
                   REGION Program funckji
                       REGION Symulacja wejsc - przepisywanie wartosci wejsciowych, gdy nie ma symulacji oprocz bWeAkt
                           IF "DB352_FF8".FF8[#i].bSt_Tryb.%X12 = 0 THEN
                               "DB352_FF8".FF8[#i].bSym.%X1 := "DB352_FF8".FF8[#i].bWeZalAuto;
                               "DB352_FF8".FF8[#i].bSym.%X8 := "DB352_FF8".FF8[#i].bWeBlZmAuto;
                               "DB352_FF8".FF8[#i].bSym.%X9 := "DB352_FF8".FF8[#i].bWeIlock;
                           END_IF;
                       END_REGION
                       REGION Okreslenie stanow
                           "DB352_FF8".FF8[#i].bSt_Tryb.%X8 := "DB352_FF8".FF8[#i].bWeAkt;
                           "DB352_FF8".FF8[#i].bSt_Tryb.%X9 := (("DB352_FF8".FF8[#i].bSym.%X8 AND "DB352_FF8".FF8[#i].bSt_Tryb.%X12) OR ("DB321_DIO".DIO[#i].bWeBlZmAuto AND NOT "DB352_FF8".FF8[#i].bSt_Tryb.%X12));
                           "DB352_FF8".FF8[#i].bSt_Tryb.%X11 := (("DB352_FF8".FF8[#i].bWeIlock AND NOT "DB352_FF8".FF8[#i].bSt_Tryb.%X12) OR ("DB352_FF8".FF8[#i].bSym.%X9 AND "DB352_FF8".FF8[#i].bSt_Tryb.%X12));
                           "DB352_FF8".FF8[#i].bSt_Tryb.%X12 := "DB352_FF8".FF8[#i].bRoZB1.%X1;
                       END_REGION
                       REGION Licznik czasu trwania impulsu
                           IF "DB352_FF8".FF8[#i].bRoZB1.%X3 AND #Imp_Sek AND NOT "DB352_FF8".FF8[#i].bPauza AND "DB352_FF8".FF8[#i].dT2_Akt=0  THEN
                               CASE "DB352_FF8".FF8[#i].iPetle OF
                                   0: "DB352_FF8".FF8[#i].dT1_old := "DB352_FF8".FF8[#i].dT1i;
                                       GOTO Warunek1;

                                   1: "DB352_FF8".FF8[#i].dT1_old := "DB352_FF8".FF8[#i].dT2i;
                                       GOTO Warunek1;

                                   2: "DB352_FF8".FF8[#i].dT1_old := "DB352_FF8".FF8[#i].dT3i;
                                       GOTO Warunek1;

                                   3: "DB352_FF8".FF8[#i].dT1_old := "DB352_FF8".FF8[#i].dT4i;
                                       GOTO Warunek1;

                                   4: "DB352_FF8".FF8[#i].dT1_old := "DB352_FF8".FF8[#i].dT5i;
                                       GOTO Warunek1;

                                   5: "DB352_FF8".FF8[#i].dT1_old := "DB352_FF8".FF8[#i].dT6i;
                                       GOTO Warunek1;

                                   6: "DB352_FF8".FF8[#i].dT1_old := "DB352_FF8".FF8[#i].dT7i;
                                       GOTO Warunek1;

                                   7: "DB352_FF8".FF8[#i].dT1_old := "DB352_FF8".FF8[#i].dT8i;
                                       GOTO Warunek1;

                                   ELSE
                                       GOTO Warunek1;
                                       ;
                               END_CASE;
                           ELSE
                               GOTO Warunek2;
                               ;
                           END_IF;
                       Warunek1:
                           "DB352_FF8".FF8[#i].dT1_Akt:="DB352_FF8".FF8[#i].dT1_Akt+1;
                           IF "DB352_FF8".FF8[#i].dT1_Akt>="DB352_FF8".FF8[#i].dT1_old THEN
                               "DB352_FF8".FF8[#i].bIhlp := 1;
                               "DB352_FF8".FF8[#i].dT1_Akt := 0;
                               "DB352_FF8".FF8[#i].iPetle := "DB352_FF8".FF8[#i].iPetle + 1;
                               ;
                           END_IF;

                           REGION Ustawianie bitu Pauzy
                           Warunek2:
                               "DB352_FF8".FF8[#i].bPauza:="DB352_FF8".FF8[#i].iPetle>="DB352_FF8".FF8[#i].iIG;
                           END_REGION
                           REGION Licznik czasu trwania przerwy miedzy impulsami
                               IF #Imp_Sek AND "DB352_FF8".FF8[#i].bRoZB1.%X3 AND NOT "DB352_FF8".FF8[#i].bPauza AND "DB352_FF8".FF8[#i].bIhlp  THEN
                                   "DB352_FF8".FF8[#i].dT2_Akt := "DB352_FF8".FF8[#i].dT2_Akt + 1;
                                   IF "DB352_FF8".FF8[#i].dT2_Akt>="DB352_FF8".FF8[#i].dT2 THEN
                                       "DB352_FF8".FF8[#i].bIhlp := 0;
                                       "DB352_FF8".FF8[#i].dT2_Akt := 0;
                                   END_IF;
                               END_IF;
                           END_REGION
                           REGION Licznik czasu trwania przerwy miedzy grupami impulsow
                               IF #Imp_Sek AND "DB352_FF8".FF8[#i].bPauza  THEN
                                   "DB352_FF8".FF8[#i].dT3_Akt := "DB352_FF8".FF8[#i].dT3_Akt + 1;
                                   IF "DB352_FF8".FF8[#i].dT3_Akt>="DB352_FF8".FF8[#i].dT3 THEN
                                       "DB352_FF8".FF8[#i].bIhlp := 0;
                                       "DB352_FF8".FF8[#i].dT3_Akt := 0;
                                       "DB352_FF8".FF8[#i].iPetle := 0;
                                   END_IF;
                               END_IF;
                           END_REGION
                           REGION Wyjscia
                               "DB352_FF8".FF8[#i].bI8 := NOT "DB352_FF8".FF8[#i].bIhlp AND "DB352_FF8".FF8[#i].iPetle = 7;

                               "DB352_FF8".FF8[#i].bI7 := NOT "DB352_FF8".FF8[#i].bIhlp AND "DB352_FF8".FF8[#i].iPetle = 6;

                               "DB352_FF8".FF8[#i].bI6 := NOT "DB352_FF8".FF8[#i].bIhlp AND "DB352_FF8".FF8[#i].iPetle = 5;

                               "DB352_FF8".FF8[#i].bI5 := NOT "DB352_FF8".FF8[#i].bIhlp AND "DB352_FF8".FF8[#i].iPetle = 4;

                               "DB352_FF8".FF8[#i].bI4 := NOT "DB352_FF8".FF8[#i].bIhlp AND "DB352_FF8".FF8[#i].iPetle = 3;

                               "DB352_FF8".FF8[#i].bI3 := NOT "DB352_FF8".FF8[#i].bIhlp AND "DB352_FF8".FF8[#i].iPetle = 2;

                               "DB352_FF8".FF8[#i].bI2 := NOT "DB352_FF8".FF8[#i].bIhlp AND "DB352_FF8".FF8[#i].iPetle = 1;

                               "DB352_FF8".FF8[#i].bI1 := NOT "DB352_FF8".FF8[#i].bIhlp AND "DB352_FF8".FF8[#i].iPetle = 0;
                           END_REGION
                           REGION Wylaczenie
                               IF NOT "DB352_FF8".FF8[#i].bRoZB1.%X3 THEN
                                   "DB352_FF8".FF8[#i].dT1_Akt := 0;
                                   "DB352_FF8".FF8[#i].dT2_Akt := 0;
                                   "DB352_FF8".FF8[#i].dT3_Akt := 0;
                                   "DB352_FF8".FF8[#i].bIhlp := 0;
                                   "DB352_FF8".FF8[#i].bI1 := 0;
                                   "DB352_FF8".FF8[#i].bI2 := 0;
                                   "DB352_FF8".FF8[#i].bI3 := 0;
                                   "DB352_FF8".FF8[#i].bI4 := 0;
                                   "DB352_FF8".FF8[#i].bI5 := 0;
                                   "DB352_FF8".FF8[#i].bI6 := 0;
                                   "DB352_FF8".FF8[#i].bI7 := 0;
                                   "DB352_FF8".FF8[#i].bI8 := 0;
                               END_IF;
                           END_REGION
                       END_REGION
                       REGION Tryb pracy i sterowanie wyjsciem
                           REGION Przepisanie potwierdzen na sterowanie reczne gdy tryb zdalny-auto
                               // Przypadek gdy ktos z wlaczonym lokalnie urz. przechodzi na tryb zdalny-reczny
                               IF "DB352_FF8".FF8[#i].bTrP=8 THEN
                                   "DB352_FF8".FF8[#i].bRoZB1.%X3 := (("DB352_FF8".FF8[#i].bWeZalAuto AND NOT "DB352_FF8".FF8[#i].bSt_Tryb.%X12) OR ("DB352_FF8".FF8[#i].bSym.%X1 AND "DB352_FF8".FF8[#i].bSt_Tryb.%X12));
                               END_IF;

                           END_REGION

                           REGION Blokada zmiany trybu zdalny-automatyczny
                               IF (("DB352_FF8".FF8[#i].bWeBlZmAuto AND NOT "DB352_FF8".FF8[#i].bSt_Tryb.%X12) OR ("DB352_FF8".FF8[#i].bSym.%X8 AND "DB352_FF8".FF8[#i].bSt_Tryb.%X12)) AND "DB352_FF8".FF8[#i].bTrP.%X3 THEN
                                   "DB352_FF8".FF8[#i].bRoZB1.%X0 := 1;
                               END_IF;
                           END_REGION
                           REGION Okreslenie trybu pracy wyjscia
                               IF "DB352_FF8".FF8[#i].bRoZB1.%X0 AND NOT "DB352_FF8".FF8[#i].bSt_Tryb.%X9 THEN
                                   "DB352_FF8".FF8[#i].bTrP := 8;
                               END_IF;
                               IF NOT "DB352_FF8".FF8[#i].bRoZB1.%X0 THEN
                                   "DB352_FF8".FF8[#i].bTrP := 4
                                   ;
                               END_IF;
                           END_REGION
                           REGION Sterowanie wyjsciem
                               "DB352_FF8".FF8[#i].bWySter := "DB352_FF8".FF8[#i].bWeZalAuto;
                           END_REGION
                           REGION Stan urzadzenia
                               IF "DB352_FF8".FF8[#i].bWySter THEN
                                   "DB352_FF8".FF8[#i].bSt_Urz := 8; //urz. wlaczone
                               ELSE
                                   "DB352_FF8".FF8[#i].bSt_Urz := 8; //urz. wylaczone
                               END_IF;
                           END_REGION
                       END_REGION
                       REGION Ustawienia koncowe
                           // Samokasowanie sygnalow
                           IF "DB352_FF8".FF8[#i].bAoff = 1 THEN
                               "DB352_FF8".FF8[#i].bWeZalAuto := 0;
                           END_IF;
                       END_REGION
                   END_REGION
               END_IF;
          END_REGION
     END_FOR;
END_FUNCTION

FUNCTION "FC353_TMR" : Void   // FC353, SCL
{ S7_Optimized_Access := 'TRUE' }
VERSION : 0.1
   VAR_INPUT
      Nr_Ost_Elementu : Int;
      Nr_Plc : Byte;
   END_VAR
   VAR_TEMP
      i : Int;
      TmrTyp : Int;
   END_VAR
BEGIN

   FOR #i := 1 TO #Nr_Ost_Elementu BY 1 DO
       REGION Opisy bitow sygnalow: bRoz,bSym,bSt,bSt_1,bTrP

           //bRoz - ROZKAZ OPERATORA - DB353.DBW10 - WORD
           //bRozB1
           //"DB353_TMR".TMR[#i].bRoZB1.%X0 - Tryb pracy: 0-Zdalny reczny; 1-Zdalny auto
           //"DB353_TMR".TMR[#i].bRoZB1.%X1 - Symulacja wejsc urz: 0-Wylaczona; 1-Zalaczona
           //"DB353_TMR".TMR[#i].bRoZB1.%X2 - Rezerwa
           //"DB353_TMR".TMR[#i].bRoZB1.%X3 - Sterowanie urz. w tr. Zdalnym-Man: 0-Wylacz; 1-Zalacz
           //"DB353_TMR".TMR[#i].bRoZB1.%X4-X7 - Rezerwa
           //
           //bRozB2 - impulsy
           //"DB353_TMR".TMR[#i].bRoZB2.%X0-X7 - Rezerwa (impuls)
           //
           //bSym - SYM WEJSCIA - DB353.DBW12 - WORD
           //"DB353_TMR".TMR[#i].bSym.%X0 - Aktywacja urz. w systemie (ustawiany tylko z programu)
           //"DB353_TMR".TMR[#i].bSym.%X1 - Sterowanie urz. w tr. Zdalnym-Auto: 0-Wylacz; 1-Zalacz
           //"DB353_TMR".TMR[#i].bSym.%X2-X7 - Rezerwa
           //"DB353_TMR".TMR[#i].bSym.%X8 - Blokada zmiany tr. zdalnego z Auto na Man: 0-Brak; 1-Aktywna
           //"DB353_TMR".TMR[#i].bSym.%X9 - Interlock w trybie Zdalnym-Auto: 0-Brak; 1-Aktywny
           //"DB353_TMR".TMR[#i].bSym.%X10-X11 - Rezerwa
           //"DB353_TMR".TMR[#i].bSym.%X12 - Zerowanie timera (kasowanie przez obiekt)
           //"DB353_TMR".TMR[#i].bSym.%X13-X15 - Rezerwa
           //
           //bSt_Tryb - STAN - DB353.DBW14 - WORD
           //"DB353_TMR".TMR[#i].bSt_Tryb.%X0-X7
           //"DB353_TMR".TMR[#i].bSt_Tryb.%X8 - Urzadzenie aktywowane
           //"DB353_TMR".TMR[#i].bSt_Tryb.%X9 - Blokada zmaiany tr. zdalnego z Auto na Man: 0-Brak; 1-Aktywna
           //"DB353_TMR".TMR[#i].bSt_Tryb.%X10 - Stan rezerwa
           //"DB353_TMR".TMR[#i].bSt_Tryb.%X11 - Interlock w trybie Zdalnym-Auto: 0-Brak; 1-Aktywny
           //"DB353_TMR".TMR[#i].bSt_Tryb.%X12 - Symulacja wejsc urzadzenia: 0-Wylaczona; 1-Zalaczona
           //"DB353_TMR".TMR[#i].bSt_Tryb.%X13 - Rezerwa
           //"DB353_TMR".TMR[#i].bSt_Tryb.%X14 - Rezerwa
           //"DB353_TMR".TMR[#i].bSt_Tryb.%X15 - Rezerwa
           //
           //bSt_Urz - STAN - DB353.DBW16 - INT
           //"DB353_TMR".TMR[#i].bSt_Urz.%X0 - STAN(1)- Awaria zbiorcza 1-Aktywna; 0-Brak aktywnosci obiektu
           //"DB353_TMR".TMR[#i].bSt_Urz.%X1 - STAN(2)- Urzadzenie: 1-Zamkniete; 0-Inny stan
           //"DB353_TMR".TMR[#i].bSt_Urz.%X2 - STAN(4)- Rezerwa
           //"DB353_TMR".TMR[#i].bSt_Urz.%X3 - STAN(8)- Urzadzenie: 1-Otwarte; 0-Inny stan
           //"DB353_TMR".TMR[#i].bSt_Urz.%X4 - STAN(16)- Rezerwa
           //"DB353_TMR".TMR[#i].bSt_Urz.%X5 - STAN(32)- Rezerwa
           //"DB353_TMR".TMR[#i].bSt_Urz.%X6-X7 - STAN(64)(128)- Rezerwa
           //
           //bTrP - TRYB PRACY - DB353.DBW17 - INT
           //"DB353_TMR".TMR[#i].bTrP.%X0 - TRYB PRACY(1) - Rezerwa
           //"DB353_TMR".TMR[#i].bTrP.%X1 - Tryb PRACY(2) - Rezerwa
           //"DB353_TMR".TMR[#i].bTrP.%X2 - TRYB PRACY(4) - Tryb Sterowania Zdalnego: 1-Zdalny Reczny; 0-Inny stan
           //"DB353_TMR".TMR[#i].bTrP.%X3 - TRYB PRACY(8) - Tryb Sterowania Zdalnego: 1-Zdalny Automatyczny; 0-Inny stan
           //"DB353_TMR".TMR[#i].bTrP.%X4-X7 - Tryb PRACY(16)(32)(64)(128) - Rezerwa
       END_REGION
       REGION Przepisanie danych do obiektu
           "DB353_TMR".TMR[#i].yNrID := #i;
           "DB353_TMR".TMR[#i].yNrPLC := #Nr_Plc;
       END_REGION
       REGION Warunek na wykonanie funkcji
           IF "DB353_TMR".TMR[#i].bWeAkt = 0 THEN //Akcja przy deaktywowaniu obiektu
               "DB353_TMR".TMR[#i].bWeAkt := 0;
               "DB353_TMR".TMR[#i].bWeZalAuto := 0;
               "DB353_TMR".TMR[#i].bWeBlZmAuto := 0;
               "DB353_TMR".TMR[#i].bWeIlock := 0;
               "DB353_TMR".TMR[#i].bWeZeruj := 0;
               "DB353_TMR".TMR[#i].bRoZB1 := 0;
               "DB353_TMR".TMR[#i].bSym := 0;
               "DB353_TMR".TMR[#i].bSt_Tryb := 0;
               "DB353_TMR".TMR[#i].bSt_Urz := 0;
               "DB353_TMR".TMR[#i].bTrP := 0;
               "DB353_TMR".TMR[#i].bWySter := 0;
           ELSE

               REGION Program funckji
                   REGION Symulacja wejsc - przepisywanie wartosci wejsciowych, gdy nie ma symulacji oprocz bWeAkt
                       IF "DB353_TMR".TMR[#i].bSt_Tryb.%X12 = 0 THEN
                           "DB353_TMR".TMR[#i].bSym.%X1 := "DB353_TMR".TMR[#i].bWeZalAuto;
                           "DB353_TMR".TMR[#i].bSym.%X8 := "DB353_TMR".TMR[#i].bWeBlZmAuto;
                           "DB353_TMR".TMR[#i].bSym.%X9 := "DB353_TMR".TMR[#i].bWeIlock;
                           "DB353_TMR".TMR[#i].bSym.%X12 := "DB353_TMR".TMR[#i].bWeZeruj;
                       END_IF;
                   END_REGION
                   REGION Okreslenie stanow
                       "DB353_TMR".TMR[#i].bSt_Tryb.%X8 := "DB353_TMR".TMR[#i].bWeAkt;
                       "DB353_TMR".TMR[#i].bSt_Tryb.%X9 := (("DB353_TMR".TMR[#i].bSym.%X8 AND "DB353_TMR".TMR[#i].bSt_Tryb.%X12) OR ("DB353_TMR".TMR[#i].bWeBlZmAuto AND NOT "DB353_TMR".TMR[#i].bSt_Tryb.%X12));
                       "DB353_TMR".TMR[#i].bSt_Tryb.%X11 := (("DB353_TMR".TMR[#i].bWeIlock AND NOT "DB353_TMR".TMR[#i].bSt_Tryb.%X12) OR ("DB353_TMR".TMR[#i].bSym.%X9 AND "DB353_TMR".TMR[#i].bSt_Tryb.%X12));
                       "DB353_TMR".TMR[#i].bSt_Tryb.%X12 := "DB353_TMR".TMR[#i].bRoZB1.%X1;
                   END_REGION
                   REGION Licznik czasu
                           IF "DB353_TMR".TMR[#i].bLatch THEN
                               #TmrTyp := 5;
                           ELSE
                               #TmrTyp := 1;
                           END_IF;

                           IF NOT "DB353_TMR".TMR[#i].bSt_Tryb.%X11 THEN
                               "FC301_Timer"(iTyp := #TmrTyp,
                                             bOnOff := ("DB353_TMR".TMR[#i].bSym.%X1 AND "DB353_TMR".TMR[#i].bSt_Tryb.%X12) OR ("DB353_TMR".TMR[#i].bWeZalAuto AND NOT "DB353_TMR".TMR[#i].bSt_Tryb.%X12),
                                             bRst := ("DB353_TMR".TMR[#i].bSym.%X12 AND "DB353_TMR".TMR[#i].bSt_Tryb.%X12) OR ("DB353_TMR".TMR[#i].bWeZeruj AND NOT "DB353_TMR".TMR[#i].bSt_Tryb.%X12),
                                             dCzasZad := "DB353_TMR".TMR[#i].dCzZad,
                                             timer_1s := "imp1s",
                                             bOk => "DB353_TMR".TMR[#i].bHlp187,
                                             dCzasAkt := "DB353_TMR".TMR[#i].dCzAkt);

                           END_IF;


                   END_REGION
                   REGION Tryb pracy i sterowanie wyjsciem
                       REGION Przepisanie potwierdzen na sterowanie reczne gdy tryb zdalny-auto
                           // Przypadek gdy ktos z wlaczonym lokalnie urz. przechodzi na tryb zdalny-reczny
                           IF "DB353_TMR".TMR[#i].bTrP = 8 THEN
                               "DB353_TMR".TMR[#i].bRoZB1.%X3 := (("DB353_TMR".TMR[#i].bWeZalAuto AND NOT "DB353_TMR".TMR[#i].bSt_Tryb.%X12) OR ("DB353_TMR".TMR[#i].bSym.%X1 AND "DB353_TMR".TMR[#i].bSt_Tryb.%X12));
                           END_IF;

                       END_REGION

                       REGION Blokada zmiany trybu zdalny-automatyczny
                           IF (("DB353_TMR".TMR[#i].bWeBlZmAuto AND NOT "DB353_TMR".TMR[#i].bSt_Tryb.%X12) OR ("DB353_TMR".TMR[#i].bSym.%X8 AND "DB353_TMR".TMR[#i].bSt_Tryb.%X12)) AND "DB353_TMR".TMR[#i].bTrP.%X3 THEN
                               "DB353_TMR".TMR[#i].bRoZB1.%X0 := 1;
                           END_IF;
                       END_REGION
                       REGION Okreslenie trybu pracy wyjscia
                           IF "DB353_TMR".TMR[#i].bRoZB1.%X0 AND NOT "DB353_TMR".TMR[#i].bSt_Tryb.%X9 THEN
                               "DB353_TMR".TMR[#i].bTrP := 8;
                           END_IF;
                           IF NOT "DB353_TMR".TMR[#i].bRoZB1.%X0 THEN
                               "DB353_TMR".TMR[#i].bTrP := 4
                               ;
                           END_IF;
                       END_REGION
                       REGION Sterowanie wyjsciem
                           "DB353_TMR".TMR[#i].bWySter := "DB353_TMR".TMR[#i].bHlp187;
                       END_REGION
                       REGION Stan urzadzenia
                           IF (("DB353_TMR".TMR[#i].bSym.%X1 AND "DB353_TMR".TMR[#i].bSt_Tryb.%X12) OR ("DB353_TMR".TMR[#i].bWeZalAuto AND NOT "DB353_TMR".TMR[#i].bSt_Tryb.%X12)) OR "DB353_TMR".TMR[#i].bWySter THEN
                               "DB353_TMR".TMR[#i].bSt_Urz := 8; //urz. wlaczone
                           ELSE
                               "DB353_TMR".TMR[#i].bSt_Urz := 2; //urz. wylaczone
                           END_IF;
                       END_REGION
                   END_REGION
                   REGION Ustawienia koncowe
                       // Samokasowanie sygnalow

                       IF ("DB353_TMR".TMR[#i].bSym.%X12 AND "DB353_TMR".TMR[#i].bSt_Tryb.%X12) OR ("DB353_TMR".TMR[#i].bWeZeruj AND NOT "DB353_TMR".TMR[#i].bSt_Tryb.%X12) THEN
                           "DB353_TMR".TMR[#i].bSym.%X12 := 0;
                           "DB353_TMR".TMR[#i].bWeZeruj := 0;
                       END_IF;

                       IF "DB353_TMR".TMR[#i].bAoff = 1 THEN
                           "DB353_TMR".TMR[#i].bWeZalAuto := 0;
                       END_IF;

                   END_REGION
               END_REGION
           END_IF;
       END_REGION
   END_FOR;
END_FUNCTION

FUNCTION "FC1000_System" : Void   // FC1000, LAD
{ S7_Optimized_Access := 'TRUE' }
VERSION : 0.1
   VAR_TEMP   // added for the SCL form of the ladder/FBD networks
      _w1 : Bool;
   END_VAR
BEGIN

REGION Network 1: Imp 1s
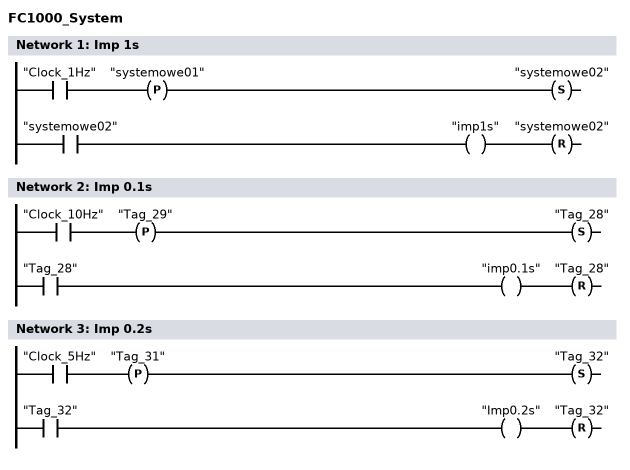
   RUNG wire#powerrail
      Contact( "Clock_1Hz" )
      P_Trig( "systemowe01" )
      S_Coil( "systemowe02" )
   END_RUNG
   RUNG wire#powerrail
      Contact( "systemowe02" )
      Coil( "imp1s" )
      R_Coil( "systemowe02" )
   END_RUNG
   // the same network as SCL:
   #_w1 := "Clock_1Hz" AND NOT "systemowe01";   // rising edge
   "systemowe01" := "Clock_1Hz";
   IF #_w1 THEN "systemowe02" := TRUE; END_IF;
   "imp1s" := "systemowe02";
   IF "systemowe02" THEN "systemowe02" := FALSE; END_IF;
END_REGION

REGION Network 2: Imp 0.1s
   RUNG wire#powerrail
      Contact( "Clock_10Hz" )
      P_Trig( "Tag_29" )
      S_Coil( "Tag_28" )
   END_RUNG
   RUNG wire#powerrail
      Contact( "Tag_28" )
      Coil( "imp0.1s" )
      R_Coil( "Tag_28" )
   END_RUNG
   // the same network as SCL:
   #_w1 := "Clock_10Hz" AND NOT "Tag_29";   // rising edge
   "Tag_29" := "Clock_10Hz";
   IF #_w1 THEN "Tag_28" := TRUE; END_IF;
   "imp0.1s" := "Tag_28";
   IF "Tag_28" THEN "Tag_28" := FALSE; END_IF;
END_REGION

REGION Network 3: Imp 0.2s
   RUNG wire#powerrail
      Contact( "Clock_5Hz" )
      P_Trig( "Tag_31" )
      S_Coil( "Tag_32" )
   END_RUNG
   RUNG wire#powerrail
      Contact( "Tag_32" )
      Coil( "Imp0.2s" )
      R_Coil( "Tag_32" )
   END_RUNG
   // the same network as SCL:
   #_w1 := "Clock_5Hz" AND NOT "Tag_31";   // rising edge
   "Tag_31" := "Clock_5Hz";
   IF #_w1 THEN "Tag_32" := TRUE; END_IF;
   "Imp0.2s" := "Tag_32";
   IF "Tag_32" THEN "Tag_32" := FALSE; END_IF;
END_REGION
END_FUNCTION

// folder: Sinamics

FUNCTION_BLOCK "DM_Objects"   // FB1, LAD
{ S7_Optimized_Access := 'TRUE' }
VERSION : 0.1
   VAR
      pump1Tank1out : "DM_Class";
      pump2Tank1in : "DM_Class";
   END_VAR
   VAR_TEMP
      i : Int;
   END_VAR
BEGIN

REGION Network 1 (SCL): Wpisanie parametrow
   #pump2Tank1in.inCircBreaker := true;
   #pump2Tank1in.inPTC := TRUE;

   #pump1Tank1out.inCircBreaker := true;
   #pump1Tank1out.inPTC := TRUE;
END_REGION

REGION Network 2: Wywolanie obiektu LAD
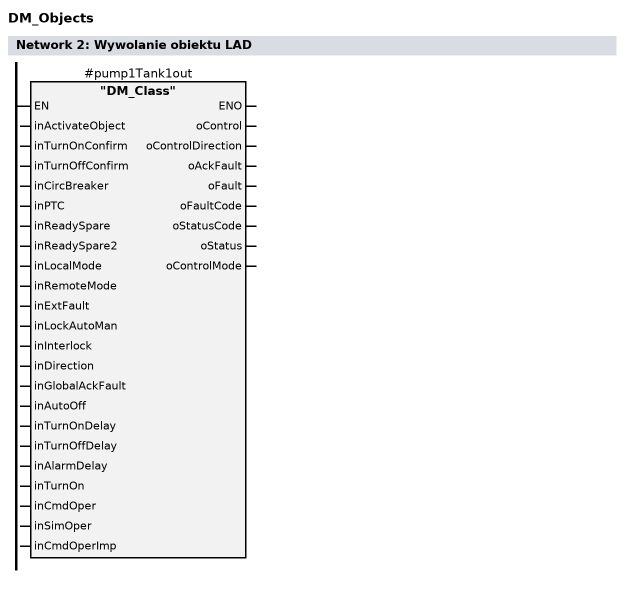
   RUNG wire#powerrail
      #pump1Tank1out(inActivateObject :=, inTurnOnConfirm :=, inTurnOffConfirm :=, inCircBreaker :=, inPTC :=, inReadySpare :=, inReadySpare2 :=, inLocalMode :=, inRemoteMode :=, inExtFault :=, inLockAutoMan :=, inInterlock :=, inDirection :=, inGlobalAckFault :=, inAutoOff :=, inTurnOnDelay :=, inTurnOffDelay :=, inAlarmDelay :=, inTurnOn :=, inCmdOper :=, inSimOper :=, inCmdOperImp :=, oControl =>, oControlDirection =>, oAckFault =>, oFault =>, oFaultCode =>, oStatusCode =>, oStatus =>, oControlMode =>)
   END_RUNG
   // the same network as SCL:
   #pump1Tank1out();   // "DM_Class"
END_REGION

REGION Network 3 (SCL): Wywolanie obiektu SCL - ladniejsze
   #pump2Tank1in();
END_REGION
END_FUNCTION_BLOCK

FUNCTION_BLOCK "DM_Sinamics"   // FB2, SCL
{ S7_Optimized_Access := 'TRUE' }
VERSION : 0.1
   VAR
      pump1Power : MC_POWER;
      pump1Control : MC_MOVEJOG;
      pump2Power : MC_POWER;
      pump2Control : MC_MOVEJOG;
   END_VAR
BEGIN

   REGION Pump 1

       #pump1Power(Axis:="pump1",
                   Enable:=NOT "DB_DM".pump1Tank1out.oFault);

       #pump1Control(Axis := "pump2",
                     JogForward := "DB_DM".pump1Tank1out.oControl AND NOT "DB_DM".pump1Tank1out.oControlDirection,
                     JogBackward := "DB_DM".pump1Tank1out.oControl AND "DB_DM".pump1Tank1out.oControlDirection);

   END_REGION


   REGION Pump 2

       #pump2Power(Axis := "pump2",
                   Enable := NOT "DB_DM".pump2Tank1in.oFault);

       #pump2Control(Axis := "pump2",
                     JogForward := "DB_DM".pump2Tank1in.oControl AND NOT "DB_DM".pump2Tank1in.oControlDirection,
                     JogBackward := "DB_DM".pump2Tank1in.oControl AND "DB_DM".pump2Tank1in.oControlDirection);

   END_REGION
END_FUNCTION_BLOCK

FUNCTION_BLOCK "DM_Class"   // FB301, SCL
{ S7_Optimized_Access := 'TRUE' }
VERSION : 0.1
   VAR_INPUT
      inActivateObject : Bool := true;   // Aktywowanie działania obiektu
      inTurnOnConfirm : Bool;   // Potwierdzenie załączenia
      inTurnOffConfirm : Bool;   // Potwierdzenie wyłączenia
      inCircBreaker : Bool;   // Gotowość obiektu - rozłącznik
      inPTC : Bool;   // Gotowość obiektu - PTC
      inReadySpare : Bool := true;   // Gotowość obiektu - rezerwa
      inReadySpare2 : Bool := true;   // Gotowość obiektu - rezerwa
      inLocalMode : Bool;   // Tryb lokalny
      inRemoteMode : Bool;   // Tryb remontowy
      inExtFault : Bool;   // Błąd zewnętrzny
      inLockAutoMan : Bool;   // Blokada przełączenia trybu Auto-Manual
      inInterlock : Bool;   // Interlok
      inDirection : Bool;   // Kierunek obrotów (1-odwrotny)
      inGlobalAckFault : Bool;   // Globalny reset
      inAutoOff : Bool;   // Resetowanie sterowania na końcu
      inTurnOnDelay : DInt;   // Czas opóźnienia załączenia [s]
      inTurnOffDelay : DInt;   // Czas opóźnienia wyłączenia [s]
      inAlarmDelay : DInt;   // Czas opóźnienia alarmu od potwierdzeń [s]
   END_VAR
   VAR_OUTPUT
      oControl : Bool;   // Wyjście sterujące
      oControlDirection : Bool;   // Wyjście strujące kierunkiem obrotów
      oAckFault : Bool;   // Wyjście reset obiektu
      oFault : Bool;   // Wyjście awaria
      oFaultCode : Byte;   // Kod awarii
      oStatusCode : Word;   // Kod statusu
      oStatus : Int;   // Status ( 1-awaria; 2-Wył; 4-Załączanie; 8-Zał; 16-Wyłączanie)
      oControlMode : Int;   // Tryb pracy (1-remont; 2-lokal; 4-manual; 8-auto)
   END_VAR
   VAR_IN_OUT
      inTurnOn : Bool;   // Załączanie z programu
      inCmdOper : Word := 16#5;   // Komendy manualne
      inSimOper : Word;   // Komendy symulacji
      inCmdOperImp : Word;   // Komendy impulsowe
   END_VAR
   VAR
      statReady : Bool;
      statManAuto : Bool;
      statSymOn : Bool;
      statSwitchEnable : Bool;
      statManTurnOn : Bool;
      statManDirection : Bool;
      statSwitchControl : Bool;
      statFaultReset : Bool;
      statActivate : Bool;
      statTurnOn : Bool;
      statTurnOnConfirm : Bool;
      statTurnOffConfirm : Bool;
      statLocal : Bool;
      statRemote : Bool;
      statExtFault : Bool;
      statLockAutoMan : Bool;
      statInterlock : Bool;
      statDirection : Bool;
      tofTurnOnDelay : TON_TIME;
      tofTurnOffDelay : TOF_TIME;
      tonAlarm : TON_TIME;
      statAlarmStart : Bool;
      statFault : Bool;
      statControlMode : Int;
      statControl : Bool;
      statTmrOnOff : Bool;
      trigGlobalReset : R_TRIG;
   END_VAR
BEGIN
   REGION Activation object - condition to execute function
       IF NOT #inActivateObject THEN
           #inTurnOn := FALSE;
           #inCmdOper := 0;
           #inSimOper := 0;
           #inCmdOperImp := 0;

           #oControl := FALSE;
           #oControlDirection := FALSE;
           #oAckFault := FALSE;
           #oFault := FALSE;
           #oFaultCode := 0;
           #oStatusCode := 0;
           #oStatus := 0;
           #oControlMode := 0;

           RETURN;

       END_IF;

   END_REGION

   REGION Rewriting inputs

       //Operator Control Word
       #statManAuto := #inCmdOper.%X0;
       #statSymOn := #inCmdOper.%X1;
       #statSwitchEnable := #inCmdOper.%X2;
       #statManTurnOn := #inCmdOper.%X3;
       #statManDirection := #inCmdOper.%X4;
       #statSwitchControl := #inCmdOper.%X6;

       //Operator Control Word Impulses
       #trigGlobalReset(CLK:=#inGlobalAckFault);

       #statFaultReset := #trigGlobalReset.Q OR #inCmdOperImp.%X0;

   END_REGION

   REGION Rewriting inputs or simulation signals to statics

       IF NOT #statSymOn THEN

           #statTurnOn := #inTurnOn;
           #statTurnOnConfirm := #inTurnOnConfirm;
           #statTurnOffConfirm := #inTurnOffConfirm;
           #statReady := #inCircBreaker AND #inPTC AND #inReadySpare AND #inReadySpare2 ;
           #statLocal := #inLocalMode;
           #statRemote := #inRemoteMode;
           #statExtFault := #inExtFault;
           #statLockAutoMan := #inLockAutoMan;
           #statInterlock := #inInterlock;
           #statDirection := #inDirection;

           //Rewriting inputs to simulation bits when simulotion is to switch fluently
           #inSimOper.%X0 := #statActivate;
           #inSimOper.%X1 := #statTurnOn;
           #inSimOper.%X2 := #statTurnOnConfirm;
           #inSimOper.%X3 := #statTurnOffConfirm;
           #inSimOper.%X4 := #statReady;
           #inSimOper.%X5 := #statLocal;
           #inSimOper.%X6 := #statRemote;
           #inSimOper.%X7 := #statExtFault;
           #inSimOper.%X8 := #statLockAutoMan;
           #inSimOper.%X9 := #statInterlock;
           #inSimOper.%X10 := #statDirection;

       ELSE

           #statActivate := #inSimOper.%X0;
           #statTurnOn := #inSimOper.%X1;
           #statTurnOnConfirm := #inSimOper.%X2;
           #statTurnOffConfirm := #inSimOper.%X3;
           #statReady:= #inSimOper.%X4;
           #statLocal := #inSimOper.%X5;
           #statRemote := #inSimOper.%X6;
           #statExtFault := #inSimOper.%X7;
           #statLockAutoMan := #inSimOper.%X8;
           #statInterlock := #inSimOper.%X9;
           #statDirection := #inSimOper.%X10;

       END_IF;


   END_REGION

   REGION Control Mode

       IF #statRemote THEN

           #statControlMode := 1;

       ELSIF #statLocal THEN

           #statControlMode := 2;

       ELSIF NOT #statManAuto AND NOT #statLockAutoMan THEN

           #statControlMode := 4;

       ELSIF #statManAuto AND NOT #statLockAutoMan THEN

           #statControlMode := 8;

       END_IF;

   END_REGION

   REGION TurnOn/Off Delay

       #tofTurnOnDelay(IN := #statTurnOn,
                       PT := 1000 * #inTurnOnDelay);

       #tofTurnOffDelay(IN := #statTurnOn,
                        PT := 1000 * #inTurnOffDelay);

       IF #tofTurnOnDelay.Q THEN

           #statTmrOnOff := TRUE;

       END_IF;

       IF NOT #tofTurnOffDelay.Q THEN

           #statTmrOnOff := FALSE;

       END_IF;
   END_REGION

   REGION Fault 
       //Zerowanie czasu awari przy zmianie sterowanie podczas ruchu - czy to w ogole cokolwiek robi???

       //Alarm from switching control 
       #statAlarmStart :=
       #statSwitchControl AND //is switch controling on
       #statSwitchEnable AND //is objects output is eneble to turn on
       #statControlMode<>2 AND //in local mode there is no alarm
       #statControlMode<>1 AND //in remote mode there is no alarm
       (
       (#statControl XOR #statTurnOnConfirm) OR //xor  0110 - if A and B have different state then =1
       (NOT #statControl XOR #statTurnOffConfirm) OR
       (#statTurnOnConfirm AND #statTurnOffConfirm) OR
       (NOT #statTurnOnConfirm AND NOT #statTurnOffConfirm)
       )
       ;
       //#tonAlarm.PT := DINT_TO_TIME(1000 * #AlarmDelay);
       //Generating switching alarm after delay
       #tonAlarm(IN := #statAlarmStart,
                 PT:=DINT_TO_TIME(1000 * #inAlarmDelay));


       //Generating fault
       IF #tonAlarm.Q OR NOT #statReady OR #statExtFault THEN

           #statFault := TRUE;

       ELSIF #statFaultReset THEN

           #statFault := FALSE;

       END_IF;

       //Fault reset 
       // IF #statFaultReset THEN
       //     #statFault := FALSE;


       // END_IF;

       //Fault code
       #oFaultCode.%X0 := #tonAlarm.Q;
       #oFaultCode.%X1 := NOT #statReady;
       #oFaultCode.%X2 := #statExtFault;
       #oFaultCode.%X3 := NOT #inCircBreaker;
       #oFaultCode.%X4 := NOT #inPTC;
       #oFaultCode.%X5 := NOT #inReadySpare;
       #oFaultCode.%X6 := NOT #inReadySpare2;

   END_REGION

   REGION Command locks

       IF #statControlMode = 8 AND #statLockAutoMan THEN

           #statManAuto := TRUE;

       ELSIF #statControlMode = 4 AND #statLockAutoMan THEN

           #statManAuto := FALSE;

       END_IF;

       // Writing states from Local to Manual when object when switching Local to Manual
       IF #statControlMode = 2 THEN

           #statManAuto := FALSE;

           IF #statTurnOffConfirm THEN

               #statTurnOn := FALSE;

           ELSIF #statTurnOnConfirm THEN

               #statTurnOn := TRUE;

           END_IF;

       END_IF;

       // Writing states from Auto to Manual when object when switching Auto to Manual
       // Przypadek gdy ktos z wlaczonym automatycznie urz. przechodzi na tryb zdalny-reczny
       IF #statControlMode = 8 THEN

           #statManTurnOn := #statTurnOn;
           #statManDirection := #statDirection;

       END_IF;

       //Resetowanie rozkazu zalaczenia w trybie manualnym po awarii
       IF #statFault THEN

           #statManTurnOn := FALSE;

       END_IF;




   END_REGION

   REGION Control output

       #statControl :=
       #statSwitchEnable AND
       NOT #statInterlock AND
       NOT #statFault AND
       ((#statControlMode = 8 AND #statTmrOnOff) OR
       (#statControlMode = 4 AND #statManTurnOn));

   END_REGION

   REGION Control Direction Output

       #oControlDirection :=
       #statSwitchEnable AND
       ((#statControlMode = 8 AND #statDirection) OR
       (#statControlMode = 4 AND #statManDirection));

   END_REGION

   REGION Reset Control

       #oAckFault := #statFaultReset;

   END_REGION ;

   REGION Device status code
       IF #statFault THEN
           #oStatus := 1;

       ELSIF #statControlMode = 1 THEN
           #oStatus := 2;

       ELSIF #statControlMode = 2 THEN

           IF #statTurnOnConfirm THEN
               #oStatus := 8;

           ELSIF #statTurnOffConfirm THEN
               #oStatus := 2;

           ELSIF #statControl THEN
               #oStatus := 4;

           ELSIF NOT #statControl THEN
               #oStatus := 16;
           END_IF;

       ELSIF #statControlMode > 2 THEN

           IF #statSwitchControl AND #statSwitchEnable THEN

               IF #statControl AND NOT #statTurnOffConfirm AND #statTurnOnConfirm THEN

                   #oStatus := 8;

               ELSIF NOT #statControl AND NOT #statTurnOnConfirm AND #statTurnOffConfirm THEN

                   #oStatus := 2;

               ELSIF #statControl THEN

                   #oStatus := 4;

               ELSIF NOT #statControl THEN

                   #oStatus := 16;

               END_IF;

           ELSIF NOT #statSwitchControl OR NOT #statSwitchEnable THEN //if no output enable or switch check then

               IF #statControl THEN

                   #oStatus := 8;

               ELSIF NOT #statControl THEN

                   #oStatus := 2;

               END_IF;

           END_IF;

       ELSE
           #oStatus := 0;

       END_IF;

   END_REGION ;


   REGION Reseting impuls
       // Samokasowanie sygnalow
       #statFaultReset := false;

       IF #inAutoOff THEN

           #statTurnOn := FALSE;

       END_IF;

   END_REGION ;

   REGION Status code


   END_REGION

   REGION Rewriting TO outputs

       #inCmdOper.%X0 := #statManAuto;
       #inCmdOper.%X1 := #statSymOn;
       #inCmdOper.%X2 := #statSwitchEnable;
       #inCmdOper.%X3 := #statManTurnOn;
       #inCmdOper.%X4 := #statManDirection;
       #inCmdOper.%X6 := #statSwitchControl;

       #inCmdOperImp.%X0 := #statFaultReset;

       #oControlMode := #statControlMode;

       #oFault := #statFault;

       #inTurnOn := #statTurnOn;

       #oControl := #statControl;
   END_REGION
END_FUNCTION_BLOCK

// ===== library types =====

// folder: LGF/4 Math operations

FUNCTION_BLOCK "LGF_Integration"   // FB10043, SCL
TITLE = LGF_Integration
{ S7_Optimized_Access := 'TRUE' }
AUTHOR : Siemens_Digital_Industries
FAMILY : LGF
NAME : LGF_Integration
// The function approximately calculates the area under a function curve. The function curve is transferred as an analog `value` (LReal) which varies over time. The integral value is output on `integral`.  
// The implementation is based on the trapezoidal rule and uses [ms] as time base.
// Diese Funktion  berechnet näherungsweise die Fläche unter einer Funktionskurve. Die Funktionskurve wird als Analogwert `value` (LReal) übergeben, der über die Zeit variiert. Am Ausgang  `integral`wird der Integralwert ausgegeben.  
// Die Implementierung beruht auf der Trapetzmethode und nutzt [ms] als Zeitbasis.
   VAR_INPUT
      enable : Bool;   // Enables integral calculation If this input is set to the value `FALSE`, the integral calculation is stopped and the `integral` output shows the last calculated value. / Aktivierung der Integral Rechnung Wird dieser Eingang auf den Wert `FALSE` berechnung gestoppt und der Ausgang `integral` zeigt den zuletzt berechneten Wert.
      value : LReal;   // Analog value of the continuous function curve, based on [ms], (e.g. [volume flow/ms]) / Analogwert der kontinuierlichen Funktionskurve, basierent auf [ms], (z.B. [Volumenstrom/ms])
      reset : Bool;   // Sets the output “integral” to “0.0”. / Setzt den Ausgang "integral" auf "0.0".
   END_VAR
   VAR_OUTPUT
      integral : LReal;   // Integral value / Integral Wert
      error : Bool;   // FALSE: No error TRUE: An error occurred during the execution of the FB / FALSE: Kein Fehler TRUE: Während der Ausführung des FB ist ein Fehler aufgetreten
      status : Word;   // 16#0000-16#7FFF: Status des FB 16#8000-16#FFFF: Fehleridentifikation (siehe folgende Tabelle) / 16#0000-16#7FFF: Status of the FB 16#8000-16#FFFF: Error identification (see following Table)
      subfunctionStatus : Word;   // Status or return value of called FB's, FC's and system blocks / Status oder Rückgabewert von aufgerufenen FB's / FC's und Systemfunktionen
   END_VAR
   VAR
      statLastTime : DTL;   // System time from previous execution of the function / Systemzeit aus dem vorhergehenden Zyklus
      statInputOldValue : LReal;   // Input value from the previous execution of the function / Eingngswert aus dem letzten vorherigem Ausführungszyklus
      statIntegral : LReal;   // Caluclated integral value / Berechneter Integral Wert
   END_VAR
   VAR_TEMP
      tempSysTime : DTL;   // Read System time / Gelesene Systemzeit
      tempTimeDiffrence : LReal;   // Time difference between the calls / Zeitdifferenz zwishcne den Funktionsaufrufen
      tempCalculation : LReal;   // Temporary variable used for passing values between calculations / Temporärer Wert um die Variablen zwischen denn Berechungen zu speichern
      tempRetval : Word;   // Return value of system function / Rückgabewert von Systemfunktonen zum Zwischenspeichern
   END_VAR
   VAR CONSTANT
      CLEAR_TIME : DTL;   // Empty DTL, to clear last saved time / Leerer DTL Datenpunkt, zum Ablöschen der Zeit
      SECOND_IN_MS : LReal := 1000.0;   // One second writen in miliseconds / Eine Sekunde in Millisekunden.
      DIVIDE_BY_TWO : LReal := 2.0;   // Constant for devision by 2 / Half the number / Konstante Zwei für Dvision / Halbierung
      ZERO : LReal := 0.0;   // Zero constant for initialization and resetting variables / Null Konstante um Variablen zu Reseten / Zurückzusetzen
      STATUS_EXECUTION_FINISHED_NO_ERROR : Word := 16#0000;   // Status: No error in the function during execution / Status: Kein Fehler während der Ausführung
      SUB_STATUS_NO_ERROR : Word := 16#0000;   // Status: No error in the called subfunction function / Status: Kein Fehler in Unterfunktions Aufrufen aufgetreten
      ERR_READ_SYS_TIME : Word := 16#8600;   // Error: System time FC `RD_SYS_T` returned an error when excuting - check `subFunctionStatus` code / Fehler: Lesen der Systemzeit `RD_SYS_T` endet mit einem Fehler - weitere infos in `subFunctionStatus`
   END_VAR
BEGIN
   REGION Block info header
     //============================================================================
     // SIEMENS AG / (c)Copyright 2017
     //----------------------------------------------------------------------------
     // Title:            LGF_Integration
     // Comment/Function: Integrates the input value
     //                   integration by trapezoidal rule
     // Library/Family:   LGF(Library General Functions)
     // Author:           Siemens Digital Industry Support
     // Tested with:      S7-PLCSIM Advanced V3.0 / S7-1215
     // Engineering:      TIA Portal V16 Update 4
     // Restrictions:     ENO disabled - no error handling by error and status
     // Requirements:     PLC (S7-1200 / S7-1500)
     //----------|------------|------------------------|----------------------------
     // Version  | Date       | Expert in charge       | Changes applied
     //----------|------------|------------------------|----------------------------
     // 01.00.00 17.02.2017  Siemens Industry Online Support
     //                      First released version
     // 01.00.01 17.08.2018  Siemens Industry Online Support
     //                      Upgrade: TIA V15 Update 2
     // 01.00.02 23.11.2018  Siemens Industry Online Support
     //                      Upgrade: TIA V15.1
     // 01.01.00 12.11.2019  Simatic Systems Support
     //                      Regions, comments and constants are added, code refactored
     // 03.00.00 23.04.2020  Simatic Systems Support
     //                      Set version to V3.0.0, harmonize the version of the whole library
     // 03.00.01 09.02.2021  Simatic Systems Support
     //                      Insert documentation
     // 03.00.02 07.06.2021  Simatic Systems Support
     //                      Fix bug - incompatibility with S7-1200 and LTIME
     //=============================================================================
   END_REGION Block info header

   REGION DESCRIPTION
     (/*NOTE
   :    The status of called commands is output in `subFunctionStatus`. In this case, the output value in `status` indicates which command caused the error. In this case, refer to the TIA Portal Online Help section for information on the respective commands.

   ---

   The integral calculation includes the summation of those trapezoidal areas that span between the last two function values on the “value” input and the time. The elapsed time is calculated via the system time of the CPU. This trapezoidal area is identical to the product of the mean value of the two process values and the time interval.

   ---

   NOTE
   :    The calculation takes [ms] as time base. So the analoge value hase to use the same time base, e.g. [volume flow/ms].

   ---

   $$
    A = \frac{1}{2} * (F_{t_1}+F_{t_0}) * (t_1-t_0) + \frac{1}{2} * (F_{t_2}+F_{t_1}) * (t_2-t_1) + ...
   $$

   Figure: Principle of operation

   ![LGF_Integration - Principle of operation](LGF_Integration.PNG "LGF_Integration - Principle of operation")

   Start the integral calculation for the inputvalue at the parameter `value`:
   * Set the parameter `enable` to the value `TRUE`
   * Set the parameter `reset` to the value `FALSE`

   If the parameter `enable` is set to the value `FALSE`, the integral calculation is stopped and the output `integral` outputs the last calculated value.  
   If the parameter `reset` is set to the value `TRUE`, the output `integral` is reset to `0.0`
   Hinweis
   :    In `subFunctionStatus` wird der Status von aufgerufenen Anweisungen ausgegeben. Der Ausgangswert in `status` gibt in diesem Fall an, welche Anweisung den Fehler verursacht hat. Holen Sie sich in diesem Fall die Informationen aus der TIA Portal Online Hilfe zu den jeweiligen Anweisungen.

   ---

   Die Integralberechnung beinhaltet die Aufsummierung jener Trapezflächen, die sich zwischen den letzten beiden Funktionswerten am Eingang "value" und der Zeit aufspannen. Die vergangene Zeit wird über die Systemzeit der CPU berechnet. Diese Trapezfläche ist identisch mit dem Produkt aus dem Mittelwert der beiden Prozesswerte und dem Zeitintervall.

   ---

   HINWEIS
   :    Die Berechnung benutzt [ms] als Zeitbasis. Das heisst, das der Analogwert die selbe Zeitbasis besitzen muss, z.B. [Volumenstrom/ms].

   ---

   $$
    A = \frac{1}{2} * (F_{t_1}+F_{t_0}) * (t_1-t_0) + \frac{1}{2} * (F_{t_2}+F_{t_1}) * (t_2-t_1) + ...
   $$

   Abbildung: Funktionsweise

   ![LGF_Integration - Funktionsweise](LGF_Integration.PNG "LGF_Integration - Funktionsweise")

   Start der Integralberechnung für den Eingangswert am Parameter `value`:  
   * Parameter `enable` auf den Wert `TRUE` setzen,
   * Parameter `reset` auf den Wert `FALSE` setzen.

   Wird der Parameter `enable` auf den Wert `FALSE` gesetzt, wird die Integralberechnung gestoppt und der Ausgang `integral` gibt den zuletzt berechneten Wert aus.  
   Wird der Parameter `reset` auf den Wert `TRUE` gesetzt, wird der Ausgang `integral` auf `0.0` zurückgesetzt.*/)
   END_REGION DESCRIPTION

   //Reset region must be before the enable region so that even if the function disabled, the user can reset the values.
   REGION Reset the function
     IF #reset THEN
       #statInputOldValue := #ZERO;
       #statIntegral := #ZERO;

       // Clear LastTime value.
       // Initial condition - first Delta time will be 0.
       #statLastTime := #CLEAR_TIME;

       #integral := #ZERO;
       #error := false;
       #status := #STATUS_EXECUTION_FINISHED_NO_ERROR;
       #subfunctionStatus := #SUB_STATUS_NO_ERROR;
       RETURN;
     END_IF;
   END_REGION Reset the function

   REGION Enable/Disable integral calculation
     IF NOT #enable THEN
       #statInputOldValue := #ZERO;

       // Clear LastTime value.
       // If it is not cleared when the function is enabled again,
       // the first value will be multiplied with the time difference of the whole disable time
       // Initial condition - first Delta time will be 0.
       #statLastTime := #CLEAR_TIME;

       #integral := #statIntegral;
       #error := false;
       #status := #STATUS_EXECUTION_FINISHED_NO_ERROR;
       #subfunctionStatus := #SUB_STATUS_NO_ERROR;
       RETURN;
     END_IF;
   END_REGION Enable/Disable integral calculation

   REGION Get system time
     // Read system time
     #tempRetval := INT_TO_WORD(RD_SYS_T(OUT => #tempSysTime));

     // Error Handling read system time
     IF (#tempRetval > #SUB_STATUS_NO_ERROR) THEN
       #integral := #statIntegral;
       #error := TRUE;
       #status := #ERR_READ_SYS_TIME;
       #subfunctionStatus := #tempRetval;
       RETURN;
     END_IF;
   END_REGION

   REGION Calculating the integral
     // Calculate time difference between last and actual time
     // coverting from DTL via time and DInt to Real
     // scale from millisecond to second
     #tempTimeDiffrence := DINT_TO_REAL(TIME_TO_DINT(T_DIFF(IN1 := #tempSysTime, IN2 := #statLastTime))) / #SECOND_IN_MS;

     // Write actual to last time
     #statLastTime := #tempSysTime;

     // integration by trapezoidal rule
     // add LastScalIn to ScalIn
     // divide by two --> avarage of both - old and actual value
     // multiply with time delta --> area unterneath the both borders
     #tempCalculation := (#value + #statInputOldValue) * #tempTimeDiffrence / #DIVIDE_BY_TWO;

     // Calculate new integral
     #statIntegral += #tempCalculation;

     // Save last input
     #statInputOldValue := #value;
   END_REGION Calculating the integral

   REGION Write outputs
     #integral := #statIntegral;
     #error := false;
     #status := #STATUS_EXECUTION_FINISHED_NO_ERROR;
     #subfunctionStatus := #SUB_STATUS_NO_ERROR;

     //ENO mechanism is not used
     ENO := TRUE;
   END_REGION Write outputs
END_FUNCTION_BLOCK

(* ===== HMI "HMI_RT_1" =====
system functions are stored by id; their names below are inferred from use
connection "HMI_Connection_1": ETHERNET, SMART_S7_1500_OMS

HMI tags "Default tag table"
   "Tag_ScreenNumber" : UInt, internal
   "Nr_AI" : Int, internal
   "Nr_AO" : Int, internal
   "Nr_DIO" : Int, internal
   "Nr_DM" : Int, internal
   "Nr_DV" : Int, internal

HMI tags "AI"
   "DB331_AI_AI{Nr}_bRoZB1" : Byte = PLC DB331_AI.AI[1].bRoZB1, 1 s
   "DB331_AI_AI{Nr}_bSym" : Word = PLC DB331_AI.AI[1].bSym AT %DB1.DBB0, 1 s
   "DB331_AI_AI{Nr}_bSt_Urz" : Int = PLC DB331_AI.AI[1].bSt_Urz AT %DB1.DBW0, 1 s
   "DB331_AI_AI{Nr}_yCzZadFiltru" : Byte = PLC DB331_AI.AI[1].yCzZadFiltru AT %DB1.DBW0, 1 s
   "DB331_AI_AI{Nr}_bB" : Byte = PLC DB331_AI.AI[1].bB AT %DB1.DBW0, 1 s
   "DB331_AI_AI{Nr}_rZH" : Real = PLC DB331_AI.AI[1].rZH AT %DB1.DBB0, 1 s
   "DB331_AI_AI{Nr}_rZL" : Real = PLC DB331_AI.AI[1].rZL AT %DB1.DBD0, 1 s
   "DB331_AI_AI{Nr}_rGHH" : Real = PLC DB331_AI.AI[1].rGHH AT %DB1.DBD0, 1 s
   "DB331_AI_AI{Nr}_rGH" : Real = PLC DB331_AI.AI[1].rGH AT %DB1.DBD0, 1 s
   "DB331_AI_AI{Nr}_rGL" : Real = PLC DB331_AI.AI[1].rGL AT %DB1.DBD0, 1 s
   "DB331_AI_AI{Nr}_rGLL" : Real = PLC DB331_AI.AI[1].rGLL AT %DB1.DBD0, 1 s
   "DB331_AI_AI{Nr}_rRoManSter" : Real = PLC DB331_AI.AI[1].rRoManSter AT %DB1.DBD0, 1 s
   "DB331_AI_AI{Nr}_rWy" : Real = PLC DB331_AI.AI[1].rWy AT %DB1.DBD0, 1 s

